
screen "Manual.Transfer" 800x480, template "TemplateWithClockAndBackBtnForManual"
   TextField "Text field_14" at 368,54 size 330x20; Text 'Cuplare contactor VFD Conveior 3 transfer palet 2'
   TextField "Text field_15" at 368,94 size 327x20; Text 'Fault Aknowledge VFD Conveior 3 transfer palet 2'
   TextField "Text field_17" at 369,134 size 267x20; Text 'ON/OFF1 VFD Conveior 3 transfer palet 2'
   TextField "Text field_18" at 369,174 size 322x20; Text 'Softstarter aer 1.1 Conveior 1 preluare paleti OK'
   TextField "Text field_19" at 369,214 size 322x20; Text 'Softstarter aer 1.2 Conveior 1 preluare paleti OK'
   TextField "Text field_20" at 369,254 size 232x20; Text 'Start Conveior 1 preluare paleti OK'
   GraphicIOField "PlotLight_Round_G" at 328,144 size 24x24; PictureOn "PilotLight_Round_G_On_256c"; PictureOff "PilotLight_Round_G_Off_256c"
      ProcessValue <- "Functionare Conveior 2 transfer palet 1"
   TextField "Text field_1" at 16,146 size 261x20; Text 'Functionare Conveior 2 transfer palet 1'
   GraphicIOField "PlotLight_Round_G_2" at 328,48 size 24x24; PictureOn "PilotLight_Round_G_On_256c"; PictureOff "PilotLight_Round_G_Off_256c"
      ProcessValue <- "Avarie Conveior 3 transfer palet 2"
   TextField "Text field_3" at 16,50 size 228x20; Text 'Avarie Conveior 3 transfer palet 2'
   GraphicIOField "PlotLight_Round_G_3" at 328,168 size 24x24; PictureOn "PilotLight_Round_G_On_256c"; PictureOff "PilotLight_Round_G_Off_256c"
      ProcessValue <- "Functionare Conveior 3 transfer palet 2"
   TextField "Text field_4" at 16,170 size 261x20; Text 'Functionare Conveior 3 transfer palet 2'
   GraphicIOField "PlotLight_Round_G_4" at 328,72 size 24x24; PictureOn "PilotLight_Round_G_On_256c"; PictureOff "PilotLight_Round_G_Off_256c"
      ProcessValue <- "Contactor cuplat Conveior 3 transfer palet 2"
   TextField "Text field_5" at 16,74 size 294x20; Text 'Contactor cuplat Conveior 3 transfer palet 2'
   GraphicIOField "PlotLight_Round_G_5" at 328,192 size 24x24; PictureOn "PilotLight_Round_G_On_256c"; PictureOff "PilotLight_Round_G_Off_256c"
      ProcessValue <- "Protectie cuplata Conveior 1 preluare paleti OK"
   TextField "Text field_6" at 16,194 size 310x20; Text 'Protectie cuplata Conveior 1 preluare paleti OK'
   GraphicIOField "PlotLight_Round_G_6" at 328,96 size 24x24; PictureOn "PilotLight_Round_G_On_256c"; PictureOff "PilotLight_Round_G_Off_256c"
      ProcessValue <- "Frana decuplata Conveior 3 transfer palet 2"
   TextField "Text field_7" at 16,98 size 289x20; Text 'Frana decuplata Conveior 3 transfer palet 2'
   GraphicIOField "PlotLight_Round_G_7" at 328,216 size 24x24; PictureOn "PilotLight_Round_G_On_256c"; PictureOff "PilotLight_Round_G_Off_256c"
      ProcessValue <- "Protectie cuplata Conveior 2 transfer palet 1"
   TextField "Text field_8" at 16,218 size 297x20; Text 'Protectie cuplata Conveior 2 transfer palet 1'
   GraphicIOField "PlotLight_Round_G_8" at 328,120 size 24x24; PictureOn "PilotLight_Round_G_On_256c"; PictureOff "PilotLight_Round_G_Off_256c"
      ProcessValue <- "Functionare Conveior 1 preluare paleti OK"
   TextField "Text field_9" at 16,122 size 274x20; Text 'Functionare Conveior 1 preluare paleti OK'
   GraphicIOField "PlotLight_Round_G_9" at 328,240 size 24x24; PictureOn "PilotLight_Round_G_On_256c"; PictureOff "PilotLight_Round_G_Off_256c"
      ProcessValue <- "Protectie cuplata Conveior 3 transfer palet 2"
   TextField "Text field_10" at 16,242 size 297x20; Text 'Protectie cuplata Conveior 3 transfer palet 2'
   Switch "Switch_2" at 696,48 size 64x32; CaptionText 'Switch'; TextOff 'OFF'; TextOn 'ON'
      on SwitchOff: ResetBit("Manual_Cuplare contactor VFD Conveior 3 transfer palet 2")
      on SwitchOn: SetBit("Manual_Cuplare contactor VFD Conveior 3 transfer palet 2")
      ProcessValue <- "Cuplare contactor VFD Conveior 3 transfer palet 2"
   Switch "Switch_5" at 697,168 size 64x32; CaptionText 'Switch'; TextOff 'OFF'; TextOn 'ON'
      on SwitchOff: ResetBit("Manual_Softstarter aer 1.1 Conveior 1 preluare paleti OK")
      on SwitchOn: SetBit("Manual_Softstarter aer 1.1 Conveior 1 preluare paleti OK")
      ProcessValue <- "Softstarter aer 1.1 Conveior 1 preluare paleti OK"
   Switch "Switch_6" at 697,208 size 64x32; CaptionText 'Switch'; TextOff 'OFF'; TextOn 'ON'
      on SwitchOff: ResetBit("Manual_Softstarter aer 1.2 Conveior 1 preluare paleti OK")
      on SwitchOn: SetBit("Manual_Softstarter aer 1.1 Conveior 1 preluare paleti OK")
      ProcessValue <- "Softstarter aer 1.2 Conveior 1 preluare paleti OK"
   TextField "Text field_2" at 369,294 size 219x20; Text 'Start Conveior 2 transfer palet 1'
   Button "DS_ACK_VFD1" at 696,90 size 73x32; TextOn 'ON'; TextOff 'OFF'
      on Release: ResetBit("Manual_Fault Aknowledge VFD Conveior 3 transfer palet 2")
      on Press: SetBit("Manual_Fault Aknowledge VFD Conveior 3 transfer palet 2")
      Appearance <- "Manual_DS_Comanda cilindru vertical jos"
   Button "DS_ON/OFF_VFD1" at 696,129 size 73x32; TextOn 'ON'; TextOff 'OFF'
      on Release: ResetBit("Manual_ON/OFF1 VFD Conveior 3 transfer palet 2")
      on Press: SetBit("Manual_ON/OFF1 VFD Conveior 3 transfer palet 2")
      Appearance <- "Manual_DS_Comanda cilindru vertical jos"
   Button "DS_ACK_VFD1_1" at 698,251 size 73x32; TextOn 'ON'; TextOff 'OFF'
      on Release: ResetBit("Manual_Start Conveior 1 preluare paleti OK")
      on Press: SetBit("Manual_Start Conveior 1 preluare paleti OK")
      Appearance <- "Manual_DS_Comanda cilindru vertical jos"
   Button "DS_ON/OFF_VFD1_1" at 698,290 size 73x32; TextOn 'ON'; TextOff 'OFF'
      on Release: ResetBit("Manual_Start Conveior 2 transfer palet 1")
      on Press: SetBit("Manual_Start Conveior 2 transfer palet 1")
      Appearance <- "Manual_DS_Comanda cilindru vertical jos"

screen "Manual.StackerBConveyors" 800x480, template "TemplateWithClockAndBackBtnForManual"
   TextField "Text field_15" at 368,54 size 296x20; Text 'Cuplare contactor VFD Conveior 1 alimentare'
   TextField "Text field_16" at 368,94 size 293x20; Text 'Fault Aknowledge VFD Conveior 1 alimentare'
   TextField "Text field_17" at 368,134 size 233x20; Text 'ON/OFF1 VFD Conveior 1 alimentare'
   TextField "Text field_18" at 368,174 size 262x20; Text 'Cuplare contactor VFD Conveior 2 iesire'
   TextField "Text field_19" at 368,214 size 259x20; Text 'Fault Aknowledge VFD Conveior 2 iesire'
   TextField "Text field_20" at 368,254 size 199x20; Text 'ON/OFF1 VFD Conveior 2 iesire'
   Switch "Switch_1" at 696,48 size 73x32; CaptionText 'Switch'; TextOff 'OFF'; TextOn 'ON'
      on SwitchOff: ResetBit("Manual_Cuplare contactor VFD Conveior 1 alimentare destacker")
      on SwitchOn: SetBit("Manual_Cuplare contactor VFD Conveior 1 alimentare destacker")
      ProcessValue <- "Manual_Cuplare contactor VFD Conveior 1 alimentare destacker"
   GraphicIOField "PlotLight_Round_G" at 280,144 size 24x24; PictureOff "PilotLight_Round_G_Off_256c"; PictureOn "PilotLight_Round_G_On_256c"
      ProcessValue <- "Protectie cuplata Conveior 1 alimentare destacker"
   TextField "Text field_1" at 16,146 size 263x20; Text 'Protectie cuplata Conveior 1 alimentare'
   GraphicIOField "PlotLight_Round_G_1" at 280,264 size 24x24; PictureOn "PilotLight_Round_G_On_256c"; PictureOff "PilotLight_Round_G_Off_256c"
      ProcessValue <- "Protectie cuplata Conveior 2 iesire destacker"
   TextField "Text field_2" at 16,266 size 229x20; Text 'Protectie cuplata Conveior 2 iesire'
   GraphicIOField "PlotLight_Round_G_2" at 280,48 size 24x24; PictureOff "PilotLight_Round_G_Off_256c"; PictureOn "PilotLight_Round_G_On_256c"
      ProcessValue <- "Avarie Conveior 1 alimentare destacker"
   TextField "Text field_3" at 16,50 size 194x20; Text 'Avarie Conveior 1 alimentare'
   GraphicIOField "PlotLight_Round_G_3" at 280,168 size 24x24; PictureOff "PilotLight_Round_G_Off_256c"; PictureOn "PilotLight_Round_G_On_256c"
      ProcessValue <- "Avarie Conveior 2 iesire destacker"
   TextField "Text field_4" at 16,170 size 160x20; Text 'Avarie Conveior 2 iesire'
   GraphicIOField "PlotLight_Round_G_4" at 280,72 size 24x24; PictureOff "PilotLight_Round_G_Off_256c"; PictureOn "PilotLight_Round_G_On_256c"
      ProcessValue <- "Contactor cuplat Conveior 1 alimentare destacker"
   TextField "Text field_5" at 16,74 size 260x20; Text 'Contactor cuplat Conveior 1 alimentare'
   GraphicIOField "PlotLight_Round_G_5" at 280,192 size 24x24; PictureOff "PilotLight_Round_G_Off_256c"; PictureOn "PilotLight_Round_G_On_256c"
      ProcessValue <- "Contactor cuplat Conveior 2 iesire destacker"
   TextField "Text field_6" at 16,194 size 226x20; Text 'Contactor cuplat Conveior 2 iesire'
   GraphicIOField "PlotLight_Round_G_6" at 280,96 size 24x24; PictureOff "PilotLight_Round_G_Off_256c"; PictureOn "PilotLight_Round_G_On_256c"
      ProcessValue <- "Frana decuplata Conveior 1 alimentare destacker"
   TextField "Text field_7" at 16,98 size 255x20; Text 'Frana decuplata Conveior 1 alimentare'
   GraphicIOField "PlotLight_Round_G_7" at 280,216 size 24x24; PictureOff "PilotLight_Round_G_Off_256c"; PictureOn "PilotLight_Round_G_On_256c"
      ProcessValue <- "Frana decuplata Conveior 2 iesire destacker"
   TextField "Text field_8" at 16,218 size 221x20; Text 'Frana decuplata Conveior 2 iesire'
   GraphicIOField "PlotLight_Round_G_8" at 280,120 size 24x24; PictureOff "PilotLight_Round_G_Off_256c"; PictureOn "PilotLight_Round_G_On_256c"
      ProcessValue <- "Functionare Conveior 1 alimentare destacker"
   TextField "Text field_9" at 16,122 size 227x20; Text 'Functionare Conveior 1 alimentare'
   GraphicIOField "PlotLight_Round_G_9" at 280,240 size 24x24; PictureOff "PilotLight_Round_G_Off_256c"; PictureOn "PilotLight_Round_G_On_256c"
      ProcessValue <- "Functionare Conveior 2 iesire destacker"
   TextField "Text field_10" at 16,242 size 193x20; Text 'Functionare Conveior 2 iesire'
   GraphicIOField "PlotLight_Round_G_10" at 280,288 size 24x24; PictureOff "PilotLight_Round_G_Off_256c"; PictureOn "PilotLight_Round_G_On_256c"
      ProcessValue <- "Senzor 1 proximitate softstarter aer destacker"
   TextField "Text field_11" at 16,290 size 243x20; Text 'Senzor 1 proximitate softstarter aer'
   GraphicIOField "PlotLight_Round_G_11" at 280,336 size 24x24; PictureOff "PilotLight_Round_G_Off_256c"; PictureOn "PilotLight_Round_G_On_256c"
      ProcessValue <- "Reset safety Stacker_New"
   TextField "Text field_12" at 16,338 size 89x20; Text 'Reset safety'
   GraphicIOField "PlotLight_Round_G_12" at 280,312 size 24x24; PictureOff "PilotLight_Round_G_Off_256c"; PictureOn "PilotLight_Round_G_On_256c"
      ProcessValue <- "Senzor 2 proximitate softstarter aer destacker"
   TextField "Text field_13" at 16,314 size 243x20; Text 'Senzor 2 proximitate softstarter aer'
   Switch "Switch_5" at 696,168 size 73x32; CaptionText 'Switch'; TextOff 'OFF'; TextOn 'ON'
      on SwitchOff: ResetBit("Manual_Cuplare contactor VFD Conveior 2 iesire destacker")
      on SwitchOn: SetBit("Manual_Cuplare contactor VFD Conveior 2 iesire destacker")
      ProcessValue <- "Manual_Cuplare contactor VFD Conveior 2 iesire destacker"
   Button "DS_ACK_VFD1" at 696,90 size 73x32; TextOn 'ON'; TextOff 'OFF'
      on Release: ResetBit("Manual_Fault Aknowledge VFD Conveior 1 alimentare destacker")
      on Press: SetBit("Manual_Fault Aknowledge VFD Conveior 1 alimentare destacker")
      Appearance <- "Manual_DS_Comanda cilindru vertical jos"
   Button "DS_ON/OFF_VFD1" at 696,129 size 73x32; TextOn 'ON'; TextOff 'OFF'
      on Release: ResetBit("Manual_ON/OFF1 VFD Conveior 1 alimentare destacker")
      on Press: SetBit("Manual_ON/OFF1 VFD Conveior 1 alimentare destacker")
      Appearance <- "Manual_DS_Comanda cilindru vertical jos"
   Button "DS_ACK_VFD2" at 696,209 size 73x32; TextOn 'ON'; TextOff 'OFF'
      on Release: ResetBit("Manual_ON/OFF1 VFD Conveior 2 iesire destacker")
      on Press: SetBit("Manual_ON/OFF1 VFD Conveior 2 iesire destacker")
      Appearance <- "Manual_DS_Comanda cilindru vertical jos"
   Button "DS_ON/OFF_VFD2" at 696,248 size 73x32; TextOn 'ON'; TextOff 'OFF'
      on Release: ResetBit("Manual_ON/OFF1 VFD Conveior 2 iesire destacker")
      on Press: SetBit("Manual_ON/OFF1 VFD Conveior 2 iesire destacker")
      Appearance <- "Manual_DS_Comanda cilindru vertical jos"

screen "Manual.StackerB" 800x480, template "TemplateWithClockAndBackBtnForManual"
   TextField "Text field_14" at 496,54 size 179x20; Text 'Comanda 1 softstarter aer'
   TextField "Text field_15" at 496,134 size 190x20; Text 'Comanda cilindru vertical jos'
   TextField "Text field_16" at 496,174 size 193x20; Text 'Comanda cilindru vertical sus'
   TextField "Text field_17" at 496,214 size 155x20; Text 'Comanda furca retrasa'
   TextField "Text field_18" at 496,254 size 153x20; Text 'Comanda furca extinsa'
   GraphicIOField "PlotLight_Round_G_2" at 160,48 size 24x24; PictureOff "PilotLight_Round_G_Off_256c"; PictureOn "PilotLight_Round_G_On_256c"
      ProcessValue <- "DB_PalletDispenser_PD2_De_Stacking_DB_PD1_MiddlePosition"
   TextField "Text field_3" at 16,50 size 126x20; Text 'PD1 MiddlePosition'
   TextField "Text field_21" at 496,94 size 179x20; Text 'Comanda 2 softstarter aer'
   GraphicIOField "PlotLight_Round_G_1" at 160,72 size 24x24; PictureOn "PilotLight_Round_G_On_256c"; PictureOff "PilotLight_Round_G_Off_256c"
      ProcessValue <- "DB_PalletDispenser_PD2_De_Stacking_DB_PD1_Up"
   TextField "Text field_1" at 16,74 size 50x20; Text 'PD1 Up'
   GraphicIOField "PlotLight_Round_G_3" at 160,96 size 24x24; PictureOn "PilotLight_Round_G_On_256c"; PictureOff "PilotLight_Round_G_Off_256c"
      ProcessValue <- "DB_PalletDispenser_PD2_De_Stacking_DB_PD1_Down"
   TextField "Text field_2" at 16,98 size 70x20; Text 'PD1 Down'
   GraphicIOField "PlotLight_Round_G_4" at 160,120 size 24x24; PictureOn "PilotLight_Round_G_On_256c"; PictureOff "PilotLight_Round_G_Off_256c"
      ProcessValue <- "DB_PalletDispenser_PD2_De_Stacking_DB_PD1_Forks_In"
   TextField "Text field_4" at 16,122 size 85x20; Text 'PD1 Forks In'
   GraphicIOField "PlotLight_Round_G_5" at 160,144 size 24x24; PictureOff "PilotLight_Round_G_Off_256c"; PictureOn "PilotLight_Round_G_On_256c"
      ProcessValue <- "DB_PalletDispenser_PD2_De_Stacking_DB_PD1_Forks_Out"
   TextField "Text field_5" at 16,146 size 95x20; Text 'PD1 Forks Out'
   GraphicIOField "PlotLight_Round_G_7" at 160,167 size 24x24; PictureOn "PilotLight_Round_G_On_256c"; PictureOff "PilotLight_Round_G_Off_256c"
      ProcessValue <- "DB_PalletDispenser_PD2_De_Stacking_DB_Alarm_Active"
   TextField "Text field_7" at 16,169 size 89x20; Text 'Alarm Active'
   GraphicIOField "PlotLight_Round_G_8" at 416,48 size 24x24; PictureOff "PilotLight_Round_G_Off_256c"; PictureOn "PilotLight_Round_G_On_256c"
      ProcessValue <- "DS_Cilindru extins"
   TextField "Text field_8" at 240,50 size 119x20; Text 'SN_Cilindru extins'
   GraphicIOField "PlotLight_Round_G_9" at 416,72 size 24x24; PictureOff "PilotLight_Round_G_Off_256c"; PictureOn "PilotLight_Round_G_On_256c"
      ProcessValue <- "DS_Cilindru retras"
   TextField "Text field_9" at 240,74 size 121x20; Text 'SN_Cilindru retras'
   GraphicIOField "PlotLight_Round_G_10" at 416,96 size 24x24; PictureOn "PilotLight_Round_G_On_256c"; PictureOff "PilotLight_Round_G_Off_256c"
      ProcessValue <- "DS_Cilindru vertical jos"
   TextField "Text field_10" at 240,98 size 152x20; Text 'SN_Cilindru vertical jos'
   GraphicIOField "PlotLight_Round_G_11" at 416,120 size 24x24; PictureOn "PilotLight_Round_G_On_256c"; PictureOff "PilotLight_Round_G_Off_256c"
      ProcessValue <- "DS_Cilindru vertical mijloc"
   TextField "Text field_11" at 240,122 size 169x20; Text 'SN_Cilindru vertical mijloc'
   GraphicIOField "PlotLight_Round_G_12" at 416,144 size 24x24; PictureOn "PilotLight_Round_G_On_256c"; PictureOff "PilotLight_Round_G_Off_256c"
      ProcessValue <- "DS_Cilindru vertical sus"
   TextField "Text field_12" at 240,146 size 155x20; Text 'SN_Cilindru vertical sus'
   GraphicIOField "PlotLight_Round_G_13" at 416,168 size 24x24; PictureOff "PilotLight_Round_G_Off_256c"; PictureOn "PilotLight_Round_G_On_256c"
      ProcessValue <- "DS_Lungime 1"
   TextField "Text field_13" at 240,170 size 94x20; Text 'SN_Lungime 1'
   GraphicIOField "PlotLight_Round_G_14" at 416,192 size 24x24; PictureOff "PilotLight_Round_G_Off_256c"; PictureOn "PilotLight_Round_G_On_256c"
      ProcessValue <- "DS_Lungime 2"
   TextField "Text field_19" at 240,194 size 94x20; Text 'SN_Lungime 2'
   GraphicIOField "PlotLight_Round_G_15" at 416,216 size 24x24; PictureOn "PilotLight_Round_G_On_256c"; PictureOff "PilotLight_Round_G_Off_256c"
      ProcessValue <- "DS_Lungime 3"
   TextField "Text field_20" at 240,218 size 94x20; Text 'SN_Lungime 3'
   GraphicIOField "PlotLight_Round_G_29" at 416,240 size 24x24; PictureOff "PilotLight_Round_G_Off_256c"; PictureOn "PilotLight_Round_G_On_256c"
      ProcessValue <- "Senzor 1 proximitate softstarter aer destacker"
   TextField "Text field_30" at 96,242 size 308x20; Text 'Senzor 1 proximitate softstarter aer stacker B'
   TextField "Text field_34" at 96,266 size 308x20; Text 'Senzor 2 proximitate softstarter aer stacker B'
   GraphicIOField "PlotLight_Round_G_33" at 416,264 size 24x24; PictureOff "PilotLight_Round_G_Off_256c"; PictureOn "PilotLight_Round_G_On_256c"
      ProcessValue <- "Senzor 2 proximitate softstarter aer destacker"
   Button "DS_Up" at 698,132 size 73x32; TextOn 'ON'; TextOff 'OFF'
      on Release: ResetBit("Manual_DS_Comanda cilindru vertical jos")
      on Press: SetBit("Manual_DS_Comanda cilindru vertical jos")
      Appearance <- "O_CilindruVerticalStacker_New_StatRet"
   Button "DS_Dwn" at 698,170 size 73x32; TextOn 'ON'; TextOff 'OFF'
      on Release: ResetBit("Manual_DS_Comanda cilindru vertical sus")
      on Press: SetBit("Manual_DS_Comanda cilindru vertical sus")
      Appearance <- "O_CilindruVerticalStacker_New_StatAv"
   Button "DS_Retr" at 698,210 size 73x32; TextOn 'ON'; TextOff 'OFF'
      on Release: ResetBit("Manual_DS_Comanda furca retrasa")
      on Press: SetBit("Manual_DS_Comanda furca retrasa")
      Appearance <- "O_FurcaStacker_New_StatRet"
   Button "DS_Av" at 698,254 size 73x32; TextOn 'ON'; TextOff 'OFF'
      on Release: ResetBit("Manual_DS_Comanda furca extinsa")
      on Press: SetBit("Manual_DS_Comanda furca extinsa")
      Appearance <- "O_FurcaStacker_New_StatAv"
   Switch "Switch_1" at 700,50 size 71x32; TextOn 'ON'; CaptionText 'Switch'; TextOff 'OFF'
      on SwitchOff: ResetBit("Manual_Comanda 1 softstarter aer destacker")
      on SwitchOn: SetBit("Manual_Comanda 1 softstarter aer destacker")
   Switch "Switch_2" at 700,88 size 71x32; TextOn 'ON'; CaptionText 'Switch'; TextOff 'OFF'
      on SwitchOn: SetBit("Manual_Comanda 2 softstarter aer destacker")
      on SwitchOff: ResetBit("Manual_Comanda 2 softstarter aer destacker")
   TextField "Text field_22" at 494,300 size 162x20; Text 'Comanda centror retras'
   TextField "Text field_23" at 494,340 size 160x20; Text 'Comanda centror extins'
   Button "S_Retr_1" at 698,296 size 73x32; TextOn 'ON'; TextOff 'OFF'
      on Release: ResetBit("O_Centror_B_ButRet")
      on Press: SetBit("O_Centror_B_ButRet")
      Appearance <- "O_Centror_B_StatRet"
   Button "S_Av_1" at 698,340 size 73x32; TextOn 'ON'; TextOff 'OFF'
      on Release: ResetBit("Manual_S_Comanda centror extins")
      on Press: SetBit("Manual_S_Comanda centror extins")
      Appearance <- "O_Centror_B_StatAv"

screen "Manual.StackerA" 800x480, template "TemplateWithClockAndBackBtnForManual"
   TextField "Text field_14" at 494,54 size 179x20; Text 'Comanda 1 softstarter aer'
   TextField "Text field_15" at 494,134 size 190x20; Text 'Comanda cilindru vertical jos'
   TextField "Text field_16" at 494,174 size 193x20; Text 'Comanda cilindru vertical sus'
   TextField "Text field_17" at 494,214 size 155x20; Text 'Comanda furca retrasa'
   TextField "Text field_18" at 494,254 size 153x20; Text 'Comanda furca extinsa'
   GraphicIOField "PlotLight_Round_G_2" at 160,48 size 24x24; PictureOn "PilotLight_Round_G_On_256c"; PictureOff "PilotLight_Round_G_Off_256c"
      ProcessValue <- "DB_PalletDispenser_PD2_Stacking_DB_PD1_MiddlePosition"
   TextField "Text field_3" at 16,50 size 126x20; Text 'PD1 MiddlePosition'
   Switch "Switch_2" at 696,48 size 64x32; CaptionText 'Switch'; TextOff 'OFF'; TextOn 'ON'
      on SwitchOff: ResetBit("Manual_Comanda 1 softstarter aer stacker")
      on SwitchOn: SetBit("Manual_Comanda 1 softstarter aer stacker")
      ProcessValue <- "Comanda 1 softstarter aer stacker"
   TextField "Text field_21" at 494,94 size 179x20; Text 'Comanda 2 softstarter aer'
   Switch "Switch_8" at 696,88 size 64x32; CaptionText 'Switch'; TextOff 'OFF'; TextOn 'ON'
      on SwitchOff: ResetBit("Manual_Comanda 2 softstarter aer stacker")
      on SwitchOn: SetBit("Manual_Comanda 2 softstarter aer stacker")
      ProcessValue <- "Comanda 2 softstarter aer stacker"
   GraphicIOField "PlotLight_Round_G_1" at 160,72 size 24x24; PictureOff "PilotLight_Round_G_Off_256c"; PictureOn "PilotLight_Round_G_On_256c"
      ProcessValue <- "DB_PalletDispenser_PD2_Stacking_DB_PD1_Up"
   TextField "Text field_1" at 16,74 size 50x20; Text 'PD1 Up'
   GraphicIOField "PlotLight_Round_G_3" at 160,96 size 24x24; PictureOff "PilotLight_Round_G_Off_256c"; PictureOn "PilotLight_Round_G_On_256c"
      ProcessValue <- "DB_PalletDispenser_PD2_Stacking_DB_PD1_Down"
   TextField "Text field_2" at 16,98 size 70x20; Text 'PD1 Down'
   GraphicIOField "PlotLight_Round_G_4" at 160,120 size 24x24; PictureOff "PilotLight_Round_G_Off_256c"; PictureOn "PilotLight_Round_G_On_256c"
      ProcessValue <- "DB_PalletDispenser_PD2_Stacking_DB_PD1_Forks_In"
   TextField "Text field_4" at 16,122 size 85x20; Text 'PD1 Forks In'
   GraphicIOField "PlotLight_Round_G_5" at 160,144 size 24x24; PictureOn "PilotLight_Round_G_On_256c"; PictureOff "PilotLight_Round_G_Off_256c"
      ProcessValue <- "DB_PalletDispenser_PD2_Stacking_DB_PD1_Forks_Out"
   TextField "Text field_5" at 16,146 size 95x20; Text 'PD1 Forks Out'
   GraphicIOField "PlotLight_Round_G_7" at 160,168 size 24x24; PictureOff "PilotLight_Round_G_Off_256c"; PictureOn "PilotLight_Round_G_On_256c"
      ProcessValue <- "DB_PalletDispenser_PD2_Stacking_DB_Alarm_Active"
   TextField "Text field_7" at 16,170 size 89x20; Text 'Alarm Active'
   GraphicIOField "PlotLight_Round_G_8" at 416,48 size 24x24; PictureOn "PilotLight_Round_G_On_256c"; PictureOff "PilotLight_Round_G_Off_256c"
      ProcessValue <- "S_Cilindru extins"
   TextField "Text field_8" at 240,50 size 111x20; Text 'S_Cilindru extins'
   GraphicIOField "PlotLight_Round_G_9" at 416,72 size 24x24; PictureOn "PilotLight_Round_G_On_256c"; PictureOff "PilotLight_Round_G_Off_256c"
      ProcessValue <- "S_Cilindru retras"
   TextField "Text field_9" at 240,74 size 113x20; Text 'S_Cilindru retras'
   GraphicIOField "PlotLight_Round_G_10" at 416,96 size 24x24; PictureOff "PilotLight_Round_G_Off_256c"; PictureOn "PilotLight_Round_G_On_256c"
      ProcessValue <- "S_Cilindru vertical jos"
   TextField "Text field_10" at 240,98 size 144x20; Text 'S_Cilindru vertical jos'
   GraphicIOField "PlotLight_Round_G_11" at 416,120 size 24x24; PictureOff "PilotLight_Round_G_Off_256c"; PictureOn "PilotLight_Round_G_On_256c"
      ProcessValue <- "S_Cilindru vertical mijloc"
   TextField "Text field_11" at 240,122 size 161x20; Text 'S_Cilindru vertical mijloc'
   GraphicIOField "PlotLight_Round_G_12" at 416,144 size 24x24; PictureOff "PilotLight_Round_G_Off_256c"; PictureOn "PilotLight_Round_G_On_256c"
      ProcessValue <- "S_Cilindru vertical sus"
   TextField "Text field_12" at 240,146 size 147x20; Text 'S_Cilindru vertical sus'
   GraphicIOField "PlotLight_Round_G_13" at 416,168 size 24x24; PictureOn "PilotLight_Round_G_On_256c"; PictureOff "PilotLight_Round_G_Off_256c"
      ProcessValue <- "S_Lungime 1"
   TextField "Text field_13" at 240,170 size 86x20; Text 'S_Lungime 1'
   GraphicIOField "PlotLight_Round_G_14" at 416,192 size 24x24; PictureOn "PilotLight_Round_G_On_256c"; PictureOff "PilotLight_Round_G_Off_256c"
      ProcessValue <- "S_Lungime 2"
   TextField "Text field_19" at 240,194 size 86x20; Text 'S_Lungime 2'
   GraphicIOField "PlotLight_Round_G_15" at 416,216 size 24x24; PictureOff "PilotLight_Round_G_Off_256c"; PictureOn "PilotLight_Round_G_On_256c"
      ProcessValue <- "S_Lungime 3"
   TextField "Text field_20" at 240,218 size 86x20; Text 'S_Lungime 3'
   GraphicIOField "PlotLight_Round_G_6" at 416,240 size 24x24; PictureOn "PilotLight_Round_G_On_256c"; PictureOff "PilotLight_Round_G_Off_256c"
      ProcessValue <- "S_Detectie palet"
   TextField "Text field_6" at 240,242 size 113x20; Text 'S_Detectie palet'
   GraphicIOField "PlotLight_Round_G_30" at 416,264 size 24x24; PictureOff "PilotLight_Round_G_Off_256c"; PictureOn "PilotLight_Round_G_On_256c"
      ProcessValue <- "Senzor 1 proximitate softstarter aer stacker"
   TextField "Text field_31" at 100,266 size 310x20; Text 'Senzor 1 proximitate softstarter aer stacker A'
   GraphicIOField "PlotLight_Round_G_34" at 416,288 size 24x24; PictureOff "PilotLight_Round_G_Off_256c"; PictureOn "PilotLight_Round_G_On_256c"
      ProcessValue <- "Senzor 2 proximitate softstarter aer stacker"
   TextField "Text field_35" at 100,290 size 310x20; Text 'Senzor 2 proximitate softstarter aer stacker A'
   Button "S_Up" at 698,132 size 73x32; TextOn 'ON'; TextOff 'OFF'
      on Release: ResetBit("Manual_S_Comanda cilindru vertical jos")
      on Press: SetBit("Manual_S_Comanda cilindru vertical jos")
      Appearance <- "O_CilindruVerticalStacker_StatRet"
   Button "S_Dwn" at 698,170 size 73x32; TextOn 'ON'; TextOff 'OFF'
      on Release: ResetBit("Manual_S_Comanda cilindru vertical sus")
      on Press: SetBit("Manual_S_Comanda cilindru vertical sus")
      Appearance <- "O_CilindruVerticalStacker_StatAv"
   Button "S_Retr" at 698,210 size 73x32; TextOn 'ON'; TextOff 'OFF'
      on Release: ResetBit("Manual_S_Comanda furca retrasa")
      on Press: SetBit("Manual_S_Comanda furca retrasa")
      Appearance <- "O_FurcaStacker_StatRet"
   Button "S_Av" at 698,254 size 73x32; TextOn 'ON'; TextOff 'OFF'
      on Release: ResetBit("Manual_S_Comanda furca extinsa")
      on Press: SetBit("Manual_S_Comanda furca extinsa")
      Appearance <- "O_FurcaStacker_StatAv"
   TextField "Text field_22" at 494,300 size 162x20; Text 'Comanda centror retras'
   TextField "Text field_23" at 494,340 size 160x20; Text 'Comanda centror extins'
   Button "S_Retr_1" at 698,296 size 73x32; TextOn 'ON'; TextOff 'OFF'
      Appearance <- "O_Centror_StatRet"
      on Press: SetBit("O_Centror_B_ButAv")
      on Release: ResetBit("O_Centror_B_ButAv")
   Button "S_Av_1" at 698,340 size 73x32; TextOn 'ON'; TextOff 'OFF'
      on Release: ResetBit("O_Centror_B_ButAv")
      on Press: SetBit("O_Centror_B_ButAv")
      Appearance <- "O_Centror_StatAv"

screen "Measurement_Error" 800x480, template "TemplateWithClockAndBackBtn"
   Button "Button_5" at 118,131 size 96x32; TextOff '1200'
      on Press: SetBit("Length_DS_HMI_1")
      Appearance <- "Fault_Length_DS"
      Visibility <- "Fault_Length_DS"
   Button "Button_6" at 118,186 size 96x32; TextOff '1600'
      on Press: SetBit("Length_DS_HMI_2")
      Appearance <- "Fault_Length_DS"
      Visibility <- "Fault_Length_DS"
   Button "Button_7" at 118,241 size 96x32; TextOff '2000'
      on Press: SetBit("Length_DS_HMI_3")
      Appearance <- "Fault_Length_DS"
      Visibility <- "Fault_Length_DS"
   Button "Button_8" at 118,296 size 96x32; TextOff 'OK'
      on Release: ResetBit("Fault_Length_DS_ACK")
      on Press: SetBit("Fault_Length_DS_ACK")
      Visibility <- "Fault_Length_DS"
   Button "Button_9" at 567,132 size 96x32; TextOff '1200'
      on Press: SetBit("Length_S_HMI_1")
      Appearance <- "Fault_Length_S"
      Visibility <- "Fault_Length_S"
   Button "Button_10" at 567,187 size 96x32; TextOff '1600'
      on Press: SetBit("Length_S_HMI_2")
      Appearance <- "Fault_Length_S"
      Visibility <- "Fault_Length_S"
   Button "Button_11" at 567,242 size 96x32; TextOff '2000'
      on Press: SetBit("Length_S_HMI_3")
      Appearance <- "Fault_Length_S"
      Visibility <- "Fault_Length_S"
   Button "Button_12" at 567,297 size 96x32; TextOff 'OK'
      on Release: ResetBit("Fault_Length_DS_ACK")
      on Press: SetBit("Fault_Length_S_ACK")
      Visibility <- "Fault_Length_S"
   TextField "Text field_1" at 68,80 size 208x42; Text 'Selectati Lungime palet Destacker'
      Visibility <- "Fault_Length_DS"
   TextField "Text field_2" at 521,80 size 188x42; Text 'Selectati Lungime palet Stacker'
      Visibility <- "Fault_Length_S"

screen "Comenzi" 800x480, template "TemplateWithClockAndBackBtn"
   Button "Button_1" at 8,392 size 136x80; TextOn 'Pagina Principala'; TextOff 'Pagina Principala'
      on Press: ActivateScreen("Main", 0)
   Switch "Switch_1" at 602,118 size 161x46; TextOn 'AUTOMAT'; CaptionText 'Switch'; TextOff 'MANUAL'
      on SwitchOff: ResetBit("Manual_DS"); SetBit("Automat_DS")
      on SwitchOn: SetBit("Manual_DS"); ResetBit("Automat_DS")
   TextField "Text field_30" at 623,83 size 112x34; Text 'Automat'
      Visibility <- "Manual_DS"
   TextField "Text field_31" at 627,83 size 97x34; Text 'Manual'
      Visibility <- "Manual_DS"
   Switch "Switch_2" at 30,106 size 160x47; TextOn 'AUTOMAT'; CaptionText 'Switch'; TextOff 'MANUAL'
      on SwitchOn: SetBit("Manual_S"); ResetBit("Automat_S")
      on SwitchOff: ResetBit("Manual_S"); SetBit("Automat_S")
   TextField "Text field_1" at 51,72 size 112x34; Text 'Automat'
      Visibility <- "Manual_S"
   TextField "Text field_2" at 55,72 size 97x34; Text 'Manual'
      Visibility <- "Manual_S"
   TextField "Text field_3" at 49,38 size 114x34; Text 'Stacking'
   TextField "Text field_4" at 602,49 size 148x34; Text 'DeStacking'
   Button "Button_2" at 58,164 size 102x37; TextOff 'Start Ciclu'
      on Press: function_b14e0dd5("bStart_S", 0)
   Button "Button_3" at 58,215 size 102x37; TextOff 'Stop Ciclu'
      on Press: function_b14e0dd5("bStop_S", 0)
   Button "Button_4" at 58,263 size 102x37; TextOff 'Pas'
      on Press: function_b14e0dd5("bStepper_S", 0)
   Button "Button_5" at 622,175 size 102x37; TextOff 'Start Ciclu'
      on Press: function_b14e0dd5("bStart_DS", 0)
   Button "Button_6" at 622,226 size 102x37; TextOff 'Stop Ciclu'
      on Press: function_b14e0dd5("bStop_SN", 0)
   Button "Button_7" at 622,274 size 102x37; TextOff 'Pas'
      on Press: function_b14e0dd5("bStepper_SN", 0)

screen "Main" 800x480, template "TemplateWithClock"
   GraphicView "Graphic view_1" at 0,21 size 800x361; Picture "Amplasament linie paleti noua_var.2"
   Button "Button_1" at 8,392 size 136x80; TextOn 'Comenzi'; TextOff 'Comenzi'
      on Press: ActivateScreen("Comenzi", 0)
   Button "Button_2" at 152,392 size 136x80; TextOff 'Mod Manual'; Authorization "Operate"
      on Press: ActivateScreen("Manual.General", 0); SetTag("CurrentScreenManual", 0)
      Visibility <- "CurrentUserGroup"
   Button "Button_3" at 296,392 size 136x80; TextOff 'Statistici Productie'; Authorization "Monitor"
      on Press: ActivateScreen("Production.Repair", 0); SetTag("CurrentScreenStatistics", 0)
      Visibility <- "CurrentUserGroup"
   Button "Button_4" at 440,392 size 136x80; TextOff 'Alarme'; Authorization "Operate"
      on Press: ActivateScreen("Alarms", 0)
   Circle "Circle_1" at 323,257 size 15x15
      Appearance <- "s_f{1}_HMI_stat_s"
   Circle "Circle_2" at 423,276 size 15x15
      Appearance <- "s_f{2}_HMI_stat_s"
   Circle "Circle_3" at 592,46 size 15x15
      Appearance <- "s_f{5}_HMI_stat_s"
   Circle "Circle_4" at 470,140 size 15x15
      Appearance <- "s_f{3}_HMI_stat_s"
   Circle "Circle_5" at 541,88 size 15x15
      Appearance <- "s_f{4}_HMI_stat_s"
   Circle "Circle_6" at 568,164 size 15x15
      Appearance <- "ds_f{1}_HMI_stat_s"
   Circle "Circle_7" at 629,116 size 15x15
      Appearance <- "ds_f{2}_HMI_stat_s"
   Circle "Circle_8" at 699,68 size 15x15
      Appearance <- "ds_f{3}_HMI_stat_s"
   GraphicView "Graphic view_10" at 370,115 size 15x15; Picture "Graphic_1"
      Visibility <- "Zone 2 112KF1 Safety Relay"
   GraphicView "Graphic view_11" at 296,216 size 15x15; Picture "Graphic_1"
      Visibility <- "Zone 2 112KF1 Safety Relay"
   GraphicView "Graphic view_12" at 545,269 size 15x15; Picture "Graphic_1"
      Visibility <- "Destacker 110KF1 Safety Relay"
   GraphicView "Graphic view_13" at 669,85 size 15x15; Picture "Graphic_1"
      Visibility <- "Destacker 111KF1 Safety Barrier Relay"
   GraphicView "Graphic view_14" at 614,181 size 15x15; Picture "Graphic_1"
      Visibility <- "Stacker 113KF1 Safety Relay"
   GraphicView "Graphic view_15" at 415,129 size 15x15; Picture "Graphic_1"
      Visibility <- "Stacker 114KF1 Safety Barrier Relay 1"
   GraphicView "Graphic view_2" at 568,61 size 15x15; Picture "Graphic_1"
      Visibility <- "Stacker 115KF1 Safety Barrier Relay 2"
   GraphicView "Graphic view_3" at 331,291 size 15x15; Picture "Graphic_1"
      Visibility <- "100KF1"
   GraphicView "Graphic view_4" at 670,196 size 15x15; Picture "Graphic_1"
      Visibility <- "Destacker 110KF1 Safety Relay"
   Group "Group_1" at 2,23 size 795x361
   AlarmView "Alarm view_1" at 0,0 size 625x23
   Button "Button_10" at 8,28 size 117x34; TextOn 'Linia A / Line A'; TextOff 'Linia A / Line A'
      on Press: SetTag("DB2_WORK_BITS_Select_MDM", 0)
      Appearance <- "DB2_WORK_BITS_Select_MDM"
   Button "Button_11" at 127,28 size 117x34; TextOn 'Linia B / Line B'; TextOff 'Linia B / Line B'
      on Press: SetTag("DB2_WORK_BITS_Select_MDM", 1)
      Appearance <- "DB2_WORK_BITS_Select_MDM"
   Button "Button_12" at 16,114 size 102x37; TextOff 'Pas'
      on Press: function_b14e0dd5("Step", 0)
   Button "Button_16" at 16,159 size 102x37; TextOff 'Stop Ciclu'
      on Press: function_b14e0dd5("Stop", 0)
   Button "Button_17" at 135,140 size 102x37; TextOn 'Automat'; TextOff 'Automat'
      on Press: SetBit("Auto"); ResetBit("Manual")
      Appearance <- "Auto"
   Button "Button_18" at 16,69 size 102x37; TextOff 'Start Ciclu'
      on Press: function_b14e0dd5("Start", 0)
   Button "Button_19" at 135,82 size 102x37; TextOn 'Manual'; TextOff 'Manual'
      on Press: SetBit("Manual"); ResetBit("Auto")
      Appearance <- "Manual"
   Rectangle "Rectangle_2" at 4,210 size 610x169
      Visibility <- "HMI.msop_viz"
   Group "Group" at 7,219 size 606x159; TextList "msjOp0"
   SymbolicIOField "Symbolic I/O field_12" at 12,219 size 595x124; TextOn '1'; TextOff '0'; TextList "msjOp0"
      Visibility <- "HMI.msop_viz"
      ProcessValue <- "pgCfg"
   Button "Button_13" at 7,344 size 167x34; TextOff 'Text'; TextList "ButOp1"
      on Press: function_b3f726e6("ButOpW", 1)
      Appearance <- "ButOpMem"
      ProcessValue <- "pgCfg"
      Visibility <- "HMI.msop_viz"
   Button "Button_14" at 226,344 size 167x34; TextOff 'Text'; TextList "ButOp2"
      on Press: function_b3f726e6("ButOpW", 2)
      Appearance <- "ButOpMem"
      ProcessValue <- "pgCfg"
      Visibility <- "HMI.msop_viz"
   Button "Button_15" at 446,344 size 167x34; TextOff 'Text'; TextList "ButOp3"
      on Press: function_b3f726e6("ButOpW", 3)
      Appearance <- "ButOpMem"
      ProcessValue <- "pgCfg"
      Visibility <- "HMI.msop_viz"
   SymbolicIOField "Symbolic I/O field_14" at 65,226 size 122x32; TextOn '1'; TextOff '0'; TextList "numeOp"
      ProcessValue <- "numSt"
      Visibility <- "HMI.msop_viz"
   SymbolicIOField "Symbolic I/O field_16" at 236,231 size 68x22; TextOn '1'; TextOff '0'; TextList "numSenz"
      ProcessValue <- "numSt"
      Visibility <- "HMI.msop_viz"
   TextField "Text field_10" at 186,233 size 51x18; Text 'Senzor:'
      Visibility <- "HMI.msop_viz"
   SymbolicIOField "Symbolic I/O field_18" at 16,226 size 51x32; TextOn '1'; TextOff '0'; TextList "loc1"
      ProcessValue <- "HMI.msop_viz"
      Visibility <- "HMI.msop_viz"
   SymbolicIOField "Symbolic I/O field_19" at 302,226 size 70x32; TextOn '1'; TextOff '0'; TextList "loc2"
      Visibility <- "HMI.msop_viz"
      ProcessValue <- "HMI.msop_viz"
   TextField "Text field_5" at 487,233 size 51x18; Text 'Senzor:'
      Visibility <- "HMI.msop_viz"
      Appearance <- "HMI.msop_viz"
   SymbolicIOField "Symbolic I/O field_15" at 371,230 size 117x25; TextOn '1'; TextOff '0'; TextList "numeOp"
      Visibility <- "HMI.msop_viz"
      ProcessValue <- "numSt_s"
      Appearance <- "HMI.msop_viz"
   SymbolicIOField "Symbolic I/O field_13" at 537,233 size 64x18; TextOn '1'; TextOff '0'; TextList "numSenz"
      Visibility <- "HMI.msop_viz"
      ProcessValue <- "numSt_s"
      Appearance <- "HMI.msop_viz"
   Line "Line_1" at 2,24 size 0x358
      Appearance <- "DB_MDM_S_step"
   Line "Line_2" at 3,23 size 388x1
      Appearance <- "DB_MDM_S_step"
   Line "Line_4" at 797,24 size 0x360
      Appearance <- "DB_MDM_SN_step"
   Line "Line_5" at 393,24 size 401x0
      Appearance <- "DB_MDM_SN_step"
   Line "Line_3" at 3,382 size 388x1
      Appearance <- "DB_MDM_S_step"
   Line "Line_6" at 393,383 size 401x0
      Appearance <- "DB_MDM_SN_step"
   Rectangle "Rectangle_1" at 185,212 size 610x169
      Visibility <- "HMI_SN_msop_vizi"
   SymbolicIOField "Symbolic I/O field_1" at 190,217 size 602x128; TextOn '1'; TextOff '0'; TextList "msjOp0"
      ProcessValue <- "pgCfg"
      Visibility <- "HMI_SN_msop_vizi"
   Button "Button_20" at 189,346 size 167x34; TextOff 'Text'; TextList "ButOp1"
      on Press: function_b3f726e6("ButOpW", 1)
      Appearance <- "ButOpMem"
      ProcessValue <- "pgCfg"
      Visibility <- "HMI_SN_msop_vizi"
   Button "Button_21" at 406,346 size 167x34; TextOff 'Text'; TextList "ButOp2"
      on Press: function_b3f726e6("ButOpW", 2)
      Appearance <- "ButOpMem"
      ProcessValue <- "pgCfg"
      Visibility <- "HMI_SN_msop_vizi"
   Button "Button_22" at 625,346 size 167x34; TextOff 'Text'; TextList "ButOp3"
      on Press: function_b3f726e6("ButOpW", 3)
      Appearance <- "ButOpMem"
      ProcessValue <- "pgCfg"
      Visibility <- "HMI_SN_msop_vizi"
   SymbolicIOField "Symbolic I/O field_2" at 244,223 size 124x32; TextOn '1'; TextOff '0'; TextList "numeOp"
      ProcessValue <- "HMI_SN_numSt"
      Visibility <- "HMI_SN_msop_vizi"
   SymbolicIOField "Symbolic I/O field_3" at 415,228 size 68x22; TextOn '1'; TextOff '0'; TextList "numSenz"
      ProcessValue <- "HMI_SN_numSt"
      Visibility <- "HMI_SN_msop_vizi"
   TextField "Text field_1" at 366,230 size 51x18; Text 'Senzor:'
      Visibility <- "HMI_SN_msop_vizi"
   SymbolicIOField "Symbolic I/O field_4" at 195,223 size 51x32; TextOn '1'; TextOff '0'; TextList "loc1"
      ProcessValue <- "HMI_SN_msop_vizi"
      Visibility <- "HMI_SN_msop_vizi"
   SymbolicIOField "Symbolic I/O field_5" at 481,223 size 70x32; TextOn '1'; TextOff '0'; TextList "loc2"
      ProcessValue <- "HMI.msop_viz"
      Visibility <- "HMI_SN_msop_vizi"
   TextField "Text field_2" at 672,230 size 51x18; Text 'Senzor:'
      Visibility <- "HMI_SN_msop_vizi"
      Appearance <- "HMI_SN_msop_vizi"
   SymbolicIOField "Symbolic I/O field_6" at 549,227 size 125x25; TextOn '1'; TextOff '0'; TextList "numeOp"
      ProcessValue <- "HMI_SN_numSt_s"
      Visibility <- "HMI_SN_msop_vizi"
      Appearance <- "HMI_SN_msop_vizi"
   SymbolicIOField "Symbolic I/O field_7" at 722,230 size 64x18; TextOn '1'; TextOff '0'; TextList "numSenz"
      Appearance <- "HMI_SN_msop_vizi"
      Visibility <- "HMI_SN_msop_vizi"
      ProcessValue <- "HMI_SN_numSt_s"

Template "TemplateWithClock" 800x480
   DateTimeField "Template_Date/time field_1" at 624,2 size 172x21
   GraphicView "Template_Graphic view_1" at 592,384 size 208x96; Picture "energom logo gonzales_1"

Template "TemplateWithClockAndBackBtn" 800x480
   Button "SB_NavigateLeft_48x48" at 72,0 size 64x40; TextOff 'Text'; PictureOff "SB_NavigateLeft_48x48_256c"
      on Press: function_efd93a16()
   Button "SB_NavigateHome_48x48" at 0,0 size 64x40; TextOff 'Text'; PictureOff "SB_NavigateHome_48x48_256c"
      on Press: ActivateScreen("Main", 0)
   DateTimeField "Template_Date/time field_1" at 624,10 size 172x21
   GraphicView "Template_Graphic view_1" at 592,384 size 208x96; Picture "energom logo gonzales_1"

Template "TemplateWithClockAndBackBtnForStatistics" 800x480
   Button "SB_NavigateHome_48x48" at 0,0 size 64x40; TextOff 'Text'; PictureOff "SB_NavigateHome_48x48_256c"
      on Press: ActivateScreen("Main", 0)
   Button "Button_4" at 8,392 size 136x80; TextOff 'Paleti Reparati'; Authorization "Operate"
      on Press: ActivateScreen("Production.Repair", 0); SetTag("CurrentScreenStatistics", 0)
      Visibility <- "CurrentUserGroup"
      Appearance <- "CurrentScreenStatistics"
   Button "Button_1" at 152,392 size 136x80; TextOff 'Paleti Demontati'; Authorization "Operate"
      on Press: ActivateScreen("Production.Destroy", 0); SetTag("CurrentScreenStatistics", 1)
      Visibility <- "CurrentUserGroup"
      Appearance <- "CurrentScreenStatistics"
   Button "Button_2" at 296,392 size 136x80; TextOff 'Energie'; Authorization "Operate"
      on Press: ActivateScreen("Energy", 0); SetTag("CurrentScreenStatistics", 2)
      Visibility <- "CurrentUserGroup"
      Appearance <- "CurrentScreenStatistics"
   Button "Button_3" at 440,392 size 136x80; TextOff 'Protectii'; Authorization "Operate"
      on Press: ActivateScreen("Safety", 0); SetTag("CurrentScreenStatistics", 3)
      Visibility <- "CurrentUserGroup"
      Appearance <- "CurrentScreenStatistics"
   DateTimeField "Template_Date/time field_1" at 624,10 size 172x21
   GraphicView "Template_Graphic view_1" at 592,384 size 208x96; Picture "energom logo gonzales_1"
   Button "Template_Button_1" at 113,5 size 53x32; TextOff 'Text'

Template "TemplateWithClockAndBackBtnForManual" 800x480
   Button "SB_NavigateHome_48x48" at 0,0 size 64x40; TextOff 'Text'; PictureOff "SB_NavigateHome_48x48_256c"
      on Press: ActivateScreen("Main", 0)
   DateTimeField "Template_Date/time field_1" at 624,10 size 172x21
   Button "Button_5" at 8,392 size 136x36; TextOff 'General'; Authorization "Operate"
      on Press: ActivateScreen("Manual.General", 0); SetTag("CurrentScreenManual", 0)
      Visibility <- "CurrentUserGroup"
      Appearance <- "CurrentScreenManual"
   Button "Button_6" at 152,392 size 136x36; TextOff 'Stacker B'; Authorization "Operate"
      on Press: ActivateScreen("Manual.StackerB", 0); SetTag("CurrentScreenManual", 2)
      Visibility <- "CurrentUserGroup"
      Appearance <- "CurrentScreenManual"
   Button "Button_7" at 296,392 size 136x36; TextOff 'Stacker A'; Authorization "Operate"
      on Press: ActivateScreen("Manual.StackerA", 0); SetTag("CurrentScreenManual", 4)
      Visibility <- "CurrentUserGroup"
      Appearance <- "CurrentScreenManual"
   Button "Button_8" at 8,436 size 136x36; TextOff 'Safety'; Authorization "Operate"
      on Press: ActivateScreen("Manual.Safety", 0); SetTag("CurrentScreenManual", 1)
      Visibility <- "CurrentUserGroup"
      Appearance <- "CurrentScreenManual"
   Button "Button_1" at 440,392 size 136x36; TextOff 'Transfer'; Authorization "Operate"
      on Press: ActivateScreen("Manual.Transfer", 0); SetTag("CurrentScreenManual", 6)
      Visibility <- "CurrentUserGroup"
      Appearance <- "CurrentScreenManual"
   GraphicView "Template_Graphic view_1" at 592,384 size 208x96; Picture "energom logo gonzales_1"
   Button "Button_2" at 152,436 size 136x36; TextOff 'Conv Stacker B'; Authorization "Operate"
      on Press: ActivateScreen("Manual.StackerBConveyors", 0); SetTag("CurrentScreenManual", 3)
      Visibility <- "CurrentUserGroup"
      Appearance <- "CurrentScreenManual"
   Button "Button_3" at 296,436 size 136x36; TextOff 'Conv Stacker A'; Authorization "Operate"
      on Press: ActivateScreen("Manual.StackerAConveyors", 0); SetTag("CurrentScreenManual", 5)
      Visibility <- "CurrentUserGroup"
      Appearance <- "CurrentScreenManual"
   Button "Button_4" at 440,436 size 136x36; TextOff 'Diagnoza IO Link'; Authorization "Operate"
      on Press: ActivateScreen("Manual.IOLinkDiag", 0); SetTag("CurrentScreenManual", 7)
      Visibility <- "CurrentUserGroup"
      Appearance <- "CurrentScreenManual"

scheduled task "ChangeUserTask"
   on Action: function_f41c6f6c("CurrentUser"); function_e1ab61de("CurrentUserGroup"); function_de9337da()
*)